AUTHOR : ISIITECH
VERSION : 0.1
// ISIITECH - Timer
// 19.01.2010 version 1.0
BEGIN

REGION Network 1 (STL): T
         A     #Input;
         JCN   ST1;
         L     #Time1;
         L     #Preset1;
         <D;
         JCN   ST2;
         A     #Pulse;
         JCN   ST2;
         L     #Time1;
         L     #Tbase;
         +D;
         T     #Time1;
         JU    ST2;
   ST1:  NOP   0;
   ST2:  NOP   0;



         A(;
         A     #RTZ;
         A     #Input_RTZ;
         );
         O(;
         AN    #Input;
         AN    #RTZ;
         );
         JCN   ST3;
         L     0;
         T     #Time1;
   ST3:  NOP   0;
END_REGION

REGION Network 2 (STL): T
         A     #Input;
         JCN   ST21;
         L     #Time2;
         L     #Preset2;
         <D;
         JCN   ST22;
         A     "point1secPls";
         JCN   ST22;
         L     #Time2;
         L     DINT#100;
         +D;
         T     #Time2;
         JU    ST22;
   ST21: NOP   0;
   ST22: NOP   0;



         A(;
         A     #RTZ;
         A     #Input_RTZ;
         );
         O(;
         AN    #Input;
         AN    #RTZ;
         );
         JCN   ST23;
         L     0;
         T     #Time2;
   ST23: NOP   0;
END_REGION
END_FUNCTION

FUNCTION "INST_CONTROL_HEATER" : Void   // FC413, LAD
TITLE = Heater controllers
{ S7_Optimized_Access := 'FALSE' }
AUTHOR : KG
VERSION : 0.1
BEGIN

REGION Network 1 (STL): Init variables
   // Dewar, Electrical Heater
         L     500.0;
         T     #Unused_TT;
         R     #ExtCmd;
END_REGION

REGION Network 2 (STL): EH90 - VB channel 1
   // Dewar, Electrical Heater
         L     2;
         T     "#DATA_HEATERS".EH90.P_TS_Ton;
         T     "#DATA_HEATERS".EH90.P_Pilot_Ton;
         L     5;
         T     "#DATA_HEATERS".EH90.P_TS_Toff;

         SET;
         A     "IOC2PLC".TT900_VALID;
         A     "EPICS_COMM_OK";
         =     #TS;
         L     "IOC2PLC".TT900;
         T     #TA;

         A(;
         L     #TA;
         L     400.0;
         >D;
         );
         JCN   _01;
         L     73.0;
         T     #TA;
   _01:  CALL  "#FC_CONTROL_HEATER"
         ( TtA      := #TA,
           TtB      := #Unused_TT,
           TtC      := #Unused_TT,
           TtD      := #Unused_TT,
           TtE      := #Unused_TT,
           TtF      := #Unused_TT,
           Nb_Tt    := 1,
           TS       := #TS,
           ExtCmd   := #ExtCmd,
           cmdEpics := "Epics_to_PLC".EH90,
           EH       := "voie 1 chaufferette BV",
           sEpics   := "PLC_to_Epics".EH90,
           Object   := "#DATA_HEATERS".EH90
         );
END_REGION

REGION Network 3 (STL): EH93-96 - VB channel 2
   // Dewar, Electrical Heater
         L     2;
         T     "#DATA_HEATERS"."EH93-96".P_TS_Ton;
         T     "#DATA_HEATERS"."EH93-96".P_Pilot_Ton;
         L     5;
         T     "#DATA_HEATERS"."EH93-96".P_TS_Toff;

         SET;
         A     "IOC2PLC".TT930_VALID;
         A     "IOC2PLC".TT940_VALID;
         A     "IOC2PLC".TT950_VALID;
         A     "IOC2PLC".TT960_VALID;
         A     "EPICS_COMM_OK";
         =     #TS;

         L     "IOC2PLC".TT930;
         T     #TA;
         A(;
         L     #TA;
         L     400.0;
         >D;
         );
         JCN   _02;
         L     73.0;
         T     #TA;
   _02:  L     "IOC2PLC".TT940;
         T     #TB;
         A(;
         L     #TB;
         L     400.0;
         >D;
         );
         JCN   _03;
         L     73.0;
         T     #TB;
   _03:  L     "IOC2PLC".TT950;
         T     #TC;
         A(;
         L     #TC;
         L     400.0;
         >D;
         );
         JCN   _04;
         L     73.0;
         T     #TC;
   _04:  L     "IOC2PLC".TT960;
         T     #TD;
         A(;
         L     #TD;
         L     400.0;
         >D;
         );
         JCN   _05;
         L     73.0;
         T     #TD;
   _05:  CALL  "#FC_CONTROL_HEATER"
         ( TtA      := #TA,
           TtB      := #TB,
           TtC      := #TC,
           TtD      := #TD,
           TtE      := #Unused_TT,
           TtF      := #Unused_TT,
           Nb_Tt    := 4,
           TS       := #TS,
           ExtCmd   := #ExtCmd,
           cmdEpics := "Epics_to_PLC"."EH93-96",
           EH       := "voie 2 chaufferette BV",
           sEpics   := "PLC_to_Epics"."EH93-96",
           Object   := "#DATA_HEATERS"."EH93-96"
         );
END_REGION

REGION Network 4 (STL): EH63_64_70 - VB channel 3
   // Dewar, Electrical Heater
         L     2;
         T     "#DATA_HEATERS"."EH63-70".P_TS_Ton;


         T     "#DATA_HEATERS"."EH63-70".P_Pilot_Ton;
         L     5;
         T     "#DATA_HEATERS"."EH63-70".P_TS_Toff;

         SET;
         A     "IOC2PLC".TT630_VALID;
         A     "IOC2PLC".TT640_VALID;
         A     "IOC2PLC".TT700_VALID;
         A     "EPICS_COMM_OK";
         =     #TS;

         CALL  "#FC_CONTROL_HEATER"
         ( TtA      := "IOC2PLC".TT630,
           TtB      := "IOC2PLC".TT640,
           TtC      := "IOC2PLC".TT700,
           TtD      := #Unused_TT,
           TtE      := #Unused_TT,
           TtF      := #Unused_TT,
           Nb_Tt    := 3,
           TS       := #TS,
           ExtCmd   := #ExtCmd,
           cmdEpics := "Epics_to_PLC"."EH63-70",
           EH       := "voie 3 chaufferette BV",
           sEpics   := "PLC_to_Epics"."EH63-70",
           Object   := "#DATA_HEATERS"."EH63-70"
         );
END_REGION

REGION Network 5 (STL): EH61-62 - VB channel 4
   // Dewar, Electrical Heater
         L     2;
         T     "#DATA_HEATERS"."EH61-62".P_TS_Ton;


         T     "#DATA_HEATERS"."EH61-62".P_Pilot_Ton;
         L     5;
         T     "#DATA_HEATERS"."EH61-62".P_TS_Toff;

         SET;
         A     "IOC2PLC".TT610_VALID;
         A     "IOC2PLC".TT620_VALID;
         A     "EPICS_COMM_OK";
         =     #TS;

         CALL  "#FC_CONTROL_HEATER"
         ( TtA      := "IOC2PLC".TT610,
           TtB      := "IOC2PLC".TT620,
           TtC      := #Unused_TT,
           TtD      := #Unused_TT,
           TtE      := #Unused_TT,
           TtF      := #Unused_TT,
           Nb_Tt    := 2,
           TS       := #TS,
           ExtCmd   := #ExtCmd,
           cmdEpics := "Epics_to_PLC"."EH61-62",
           EH       := "voie 4 chaufferette BV",
           sEpics   := "PLC_to_Epics"."EH61-62",
           Object   := "#DATA_HEATERS"."EH61-62"
         );
END_REGION

REGION Network 6 (STL): EH60_67-69 - VB channel 5
   // Dewar, Electrical Heater
         L     2;
         T     "#DATA_HEATERS"."EH60_67-69".P_TS_Ton;


         T     "#DATA_HEATERS"."EH60_67-69".P_Pilot_Ton;
         L     5;
         T     "#DATA_HEATERS"."EH60_67-69".P_TS_Toff;

         SET;
         A     "IOC2PLC".TT600_VALID;
         A     "IOC2PLC".TT670_VALID;
         A     "IOC2PLC".TT680_VALID;
         A     "IOC2PLC".TT690_VALID;
         A     "EPICS_COMM_OK";
         =     #TS;

         CALL  "#FC_CONTROL_HEATER"
         ( TtA      := "IOC2PLC".TT600,
           TtB      := "IOC2PLC".TT670,
           TtC      := "IOC2PLC".TT680,
           TtD      := "IOC2PLC".TT690,
           TtE      := #Unused_TT,
           TtF      := #Unused_TT,
           Nb_Tt    := 4,
           TS       := #TS,
           ExtCmd   := #ExtCmd,
           cmdEpics := "Epics_to_PLC"."EH60_67-69",
           EH       := "voie 5 chaufferette BV",
           sEpics   := "PLC_to_Epics"."EH60_67-69",
           Object   := "#DATA_HEATERS"."EH60_67-69"
         );
END_REGION

REGION Network 7 (STL): EH97-98 - VB channel 6
   // Dewar, Electrical Heater
         L     2;
         T     "#DATA_HEATERS"."EH97-98".P_TS_Ton;
         T     "#DATA_HEATERS"."EH97-98".P_Pilot_Ton;
         L     5;
         T     "#DATA_HEATERS"."EH97-98".P_TS_Toff;

         SET;
         A     "IOC2PLC".TT970_VALID;
         A     "IOC2PLC".TT980_VALID;
         A     "EPICS_COMM_OK";
         =     #TS;

         L     "IOC2PLC".TT970;
         T     #TA;
         A(;
         L     #TA;
         L     400.0;
         >D;
         );
         JCN   _61;
         L     73.0;
         T     #TA;
   _61:  L     "IOC2PLC".TT980;
         T     #TB;
         A(;
         L     #TB;
         L     400.0;
         >D;
         );
         JCN   _62;
         L     73.0;
         T     #TB;

   _62:  CALL  "#FC_CONTROL_HEATER"
         ( TtA      := #TA,
           TtB      := #TB,
           TtC      := #Unused_TT,
           TtD      := #Unused_TT,
           TtE      := #Unused_TT,
           TtF      := #Unused_TT,
           Nb_Tt    := 2,
           TS       := #TS,
           ExtCmd   := #ExtCmd,
           cmdEpics := "Epics_to_PLC"."EH97-98",
           EH       := "voie 6 chaufferette BV",
           sEpics   := "PLC_to_Epics"."EH97-98",
           Object   := "#DATA_HEATERS"."EH97-98"
         );
END_REGION

REGION Network 8 (STL): EH903 - CM channel 2
   // Dewar, Electrical Heater
         L     2;
         T     "#DATA_HEATERS".EH903.P_TS_Ton;
         T     "#DATA_HEATERS".EH903.P_Pilot_Ton;
         L     5;
         T     "#DATA_HEATERS".EH903.P_TS_Toff;

         SET;
         A     "IOC2PLC".TT903_VALID;
         A     "EPICS_COMM_OK";
         =     #TS;

         L     "IOC2PLC".TT903;
         T     #TA;
         A(;
         L     #TA;
         L     400.0;
         >D;
         );
         JCN   _121;
         L     73.0;
         T     #TA;
   _121: CALL  "#FC_CONTROL_HEATER"
         ( TtA      := #TA,
           TtB      := #Unused_TT,
           TtC      := #Unused_TT,
           TtD      := #Unused_TT,
           TtE      := #Unused_TT,
           TtF      := #Unused_TT,
           Nb_Tt    := 1,
           TS       := #TS,
           ExtCmd   := #ExtCmd,
           cmdEpics := "Epics_to_PLC".EH903,
           EH       := "voie 2 chaufferette CM",
           sEpics   := "PLC_to_Epics".EH903,
           Object   := "#DATA_HEATERS".EH903
         );
END_REGION

REGION Network 9 (STL): EH920 - CM channel 3
   // Dewar, Electrical Heater
         L     2;
         T     "#DATA_HEATERS".EH920.P_TS_Ton;
         T     "#DATA_HEATERS".EH920.P_Pilot_Ton;
         L     5;
         T     "#DATA_HEATERS".EH920.P_TS_Toff;

         SET;
         A     "IOC2PLC".TT920_CM_VALID;
         A     "EPICS_COMM_OK";
         =     #TS;

         L     "IOC2PLC".TT920_CM;
         T     #TA;
         A(;
         L     #TA;
         L     400.0;
         >D;
         );
         JCN   _131;
         L     73.0;
         T     #TA;
   _131: CALL  "#FC_CONTROL_HEATER"
         ( TtA      := #TA,
           TtB      := #Unused_TT,
           TtC      := #Unused_TT,
           TtD      := #Unused_TT,
           TtE      := #Unused_TT,
           TtF      := #Unused_TT,
           Nb_Tt    := 1,
           TS       := #TS,
           ExtCmd   := #ExtCmd,
           cmdEpics := "Epics_to_PLC".EH920,
           EH       := "voie 3 chaufferette CM",
           sEpics   := "PLC_to_Epics".EH920,
           Object   := "#DATA_HEATERS".EH920
         );
END_REGION

REGION Network 10 (STL): EH918 - CM channel 9
   // Dewar, Electrical Heater
         L     2;
         T     "#DATA_HEATERS".EH918.P_TS_Ton;
         T     "#DATA_HEATERS".EH918.P_Pilot_Ton;
         L     5;
         T     "#DATA_HEATERS".EH918.P_TS_Toff;

         SET;
         A     "IOC2PLC".TT918_VALID;
         A     "EPICS_COMM_OK";
         =     #TS;

         L     "IOC2PLC".TT918;
         T     #TA;
         A(;
         L     #TA;
         L     400.0;
         >D;
         );
         JCN   _191;
         L     73.0;
         T     #TA;
   _191: CALL  "#FC_CONTROL_HEATER"
         ( TtA      := #TA,
           TtB      := #Unused_TT,
           TtC      := #Unused_TT,
           TtD      := #Unused_TT,
           TtE      := #Unused_TT,
           TtF      := #Unused_TT,
           Nb_Tt    := 1,
           TS       := #TS,
           ExtCmd   := #ExtCmd,
           cmdEpics := "Epics_to_PLC".EH918,
           EH       := "voie 9 chaufferette CM",
           sEpics   := "PLC_to_Epics".EH918,
           Object   := "#DATA_HEATERS".EH918
         );
END_REGION

REGION Network 11 (STL): EH904 - CM channel 11
   // Dewar, Electrical Heater
         L     2;
         T     "#DATA_HEATERS".EH904.P_TS_Ton;
         T     "#DATA_HEATERS".EH904.P_Pilot_Ton;
         L     5;
         T     "#DATA_HEATERS".EH904.P_TS_Toff;

         SET;
         A     "IOC2PLC".TT904_VALID;
         A     "EPICS_COMM_OK";
         =     #TS;

         L     "IOC2PLC".TT904;
         T     #TA;
         A(;
         L     #TA;
         L     400.0;
         >D;
         );
         JCN   _1111;
         L     73.0;
         T     #TA;
   _1111:CALL  "#FC_CONTROL_HEATER"
         ( TtA      := #TA,
           TtB      := #Unused_TT,
           TtC      := #Unused_TT,
           TtD      := #Unused_TT,
           TtE      := #Unused_TT,
           TtF      := #Unused_TT,
           Nb_Tt    := 1,
           TS       := #TS,
           ExtCmd   := #ExtCmd,
           cmdEpics := "Epics_to_PLC".EH904,
           EH       := "voie 11 chaufferette CM",
           sEpics   := "PLC_to_Epics".EH904,
           Object   := "#DATA_HEATERS".EH904
         );
END_REGION

REGION Network 12 (STL): EH13 - Coupler 1 flange
   // Dewar, Electrical Heater
         L     2;
         T     "#DATA_HEATERS".EH13.P_TS_Ton;
         T     "#DATA_HEATERS".EH13.P_Pilot_Ton;
         L     5;
         T     "#DATA_HEATERS".EH13.P_TS_Toff;

         L     "PLC_to_Epics".TT103.Visu;
         L     0;
         ==I;
         =     #Enable;
         CALL  "#FC_CONTROL_HEATER"
         ( TtA      := "PLC_to_Epics".TT103.Level,
           TtB      := #Unused_TT,
           TtC      := #Unused_TT,
           TtD      := #Unused_TT,
           TtE      := #Unused_TT,
           TtF      := #Unused_TT,
           Nb_Tt    := 1,
           TS       := #Enable,
           ExtCmd   := #ExtCmd,
           cmdEpics := "Epics_to_PLC".EH13,
           EH       := "EH13 Cpl1",
           sEpics   := "PLC_to_Epics".EH13,
           Object   := "#DATA_HEATERS".EH13
         );
END_REGION

REGION Network 13 (STL): EH43 - Coupler 2 flange
   // Dewar, Electrical Heater
         L     2;
         T     "#DATA_HEATERS".EH43.P_TS_Ton;
         T     "#DATA_HEATERS".EH43.P_Pilot_Ton;
         L     5;
         T     "#DATA_HEATERS".EH43.P_TS_Toff;

         L     "PLC_to_Epics".TT203.Visu;
         L     0;
         ==I;
         =     #Enable;
         CALL  "#FC_CONTROL_HEATER"
         ( TtA      := "PLC_to_Epics".TT203.Level,
           TtB      := #Unused_TT,
           TtC      := #Unused_TT,
           TtD      := #Unused_TT,
           TtE      := #Unused_TT,
           TtF      := #Unused_TT,
           Nb_Tt    := 1,
           TS       := #Enable,
           ExtCmd   := #ExtCmd,
           cmdEpics := "Epics_to_PLC".EH43,
           EH       := "EH43 Cpl2",
           sEpics   := "PLC_to_Epics".EH43,
           Object   := "#DATA_HEATERS".EH43
         );
END_REGION
END_FUNCTION

FUNCTION "Manage_HEATERS" : Void   // FC513, LAD
TITLE = Manage the heaters
{ S7_Optimized_Access := 'FALSE' }
AUTHOR : KG
VERSION : 0.1
BEGIN

REGION Network 1: EH13 & EH43 - Coupler flange cavity 1 and 2
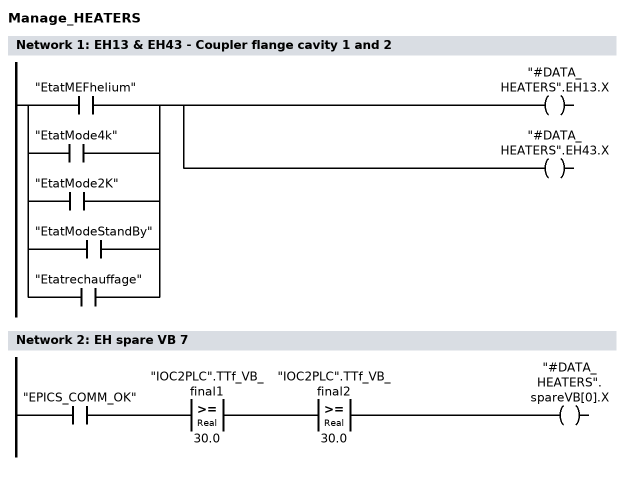
   RUNG wire#powerrail
      Contact( "EtatMEFhelium" )
      wire#w1
      Coil( "#DATA_HEATERS".EH13.X )
   END_RUNG
   RUNG wire#powerrail
      Contact( "EtatMode4k" )
   END_RUNG wire#w1
   RUNG wire#powerrail
      Contact( "EtatMode2K" )
   END_RUNG wire#w1
   RUNG wire#powerrail
      Contact( "EtatModeStandBy" )
   END_RUNG wire#w1
   RUNG wire#powerrail
      Contact( "Etatrechauffage" )
   END_RUNG wire#w1
   RUNG wire#w1
      Coil( "#DATA_HEATERS".EH43.X )
   END_RUNG
   // the same network as SCL:
   "#DATA_HEATERS".EH13.X := "EtatMEFhelium" OR "EtatMode4k" OR "EtatMode2K" OR "EtatModeStandBy" OR "Etatrechauffage";
   "#DATA_HEATERS".EH43.X := "#DATA_HEATERS".EH13.X;
END_REGION

REGION Network 2: EH spare VB 7
   RUNG wire#powerrail
      Contact( "EPICS_COMM_OK" )
      { S7_Templates := "SrcType := Real" } GE_Contact(in1 := "IOC2PLC".TTf_VB_final1, in2 := 30.0)
      { S7_Templates := "SrcType := Real" } GE_Contact(in1 := "IOC2PLC".TTf_VB_final2, in2 := 30.0)
      Coil( "#DATA_HEATERS".spareVB[0].X )
   END_RUNG
   // the same network as SCL:
   "#DATA_HEATERS".spareVB[0].X := "EPICS_COMM_OK" AND ("IOC2PLC".TTf_VB_final1 >= 30.0) AND ("IOC2PLC".TTf_VB_final2 >= 30.0);
END_REGION
END_FUNCTION

ORGANIZATION_BLOCK "Main"   // OB1, STL
TITLE = "Main Program Sweep (Cycle)"
{ S7_Optimized_Access := 'FALSE' }
VERSION : 0.1
BEGIN

REGION Network 1: Set-up the timing pulse for FC_TIMER
         A     "point1sec";
         AN    "point1secMem";
         =     "point1secPls";
         A     "point1sec";
         =     "point1secMem";

         SET;
         A     "oneSec";
         AN    "oneSecMem";
         =     "oneSecPls";
         A     "oneSec";
         =     "oneSecMem";
END_REGION

REGION Network 2: Get data and commands from Epics IOC
         CALL  "Recv_from_Epics";
         NOP   0;
END_REGION

REGION Network 3
         A     "Graph/manuelle";
         JNB   Label_0;
         CALL  "commande vanne";
   Label_0:NOP   0;
END_REGION

REGION Network 4
         CALL  "NIveau Helium&Pression&vide";
         NOP   0;
END_REGION

REGION Network 5
         CALL  "ACQ_CABTF";
         NOP   0;
END_REGION

REGION Network 6
         AN    "Graph/manuelle";
         JNB   Label_1;
         CALL  "grafcet";
   Label_1:NOP   0;
END_REGION

REGION Network 7
         CALL  "Send_to_Epics";
         NOP   0;
END_REGION

REGION Network 8: Instantiate the heaters control
         CALL  "INST_CONTROL_HEATER";
END_REGION

REGION Network 9: Manage the heaters
         CALL  "Manage_HEATERS";
END_REGION

REGION Network 10: Clear INIT flag after the first cycle
         SET;
         R     "INIT";
END_REGION

REGION Network 11
         CALL  "UpdateData2HNOSS";
END_REGION

REGION Network 12: Appeler le bloc de diagnostic système / Call system diagnostics block
         CALL  "RSE_FB", "RSE_DB";
END_REGION
END_ORGANIZATION_BLOCK

ORGANIZATION_BLOCK "CYC_INT2"   // OB32, LAD
TITLE = Cyclic_1s / "Cyclic Interrupt"
{ S7_Optimized_Access := 'FALSE' }
AUTHOR : KG
VERSION : 0.1
// Call the PID functionswith 1s interval
   VAR_TEMP   // added for the SCL form of the ladder/FBD networks
      _w1 : Bool;
   END_VAR
BEGIN

REGION Network 1: PID regulator for the LN2 screen cooling (CV60)
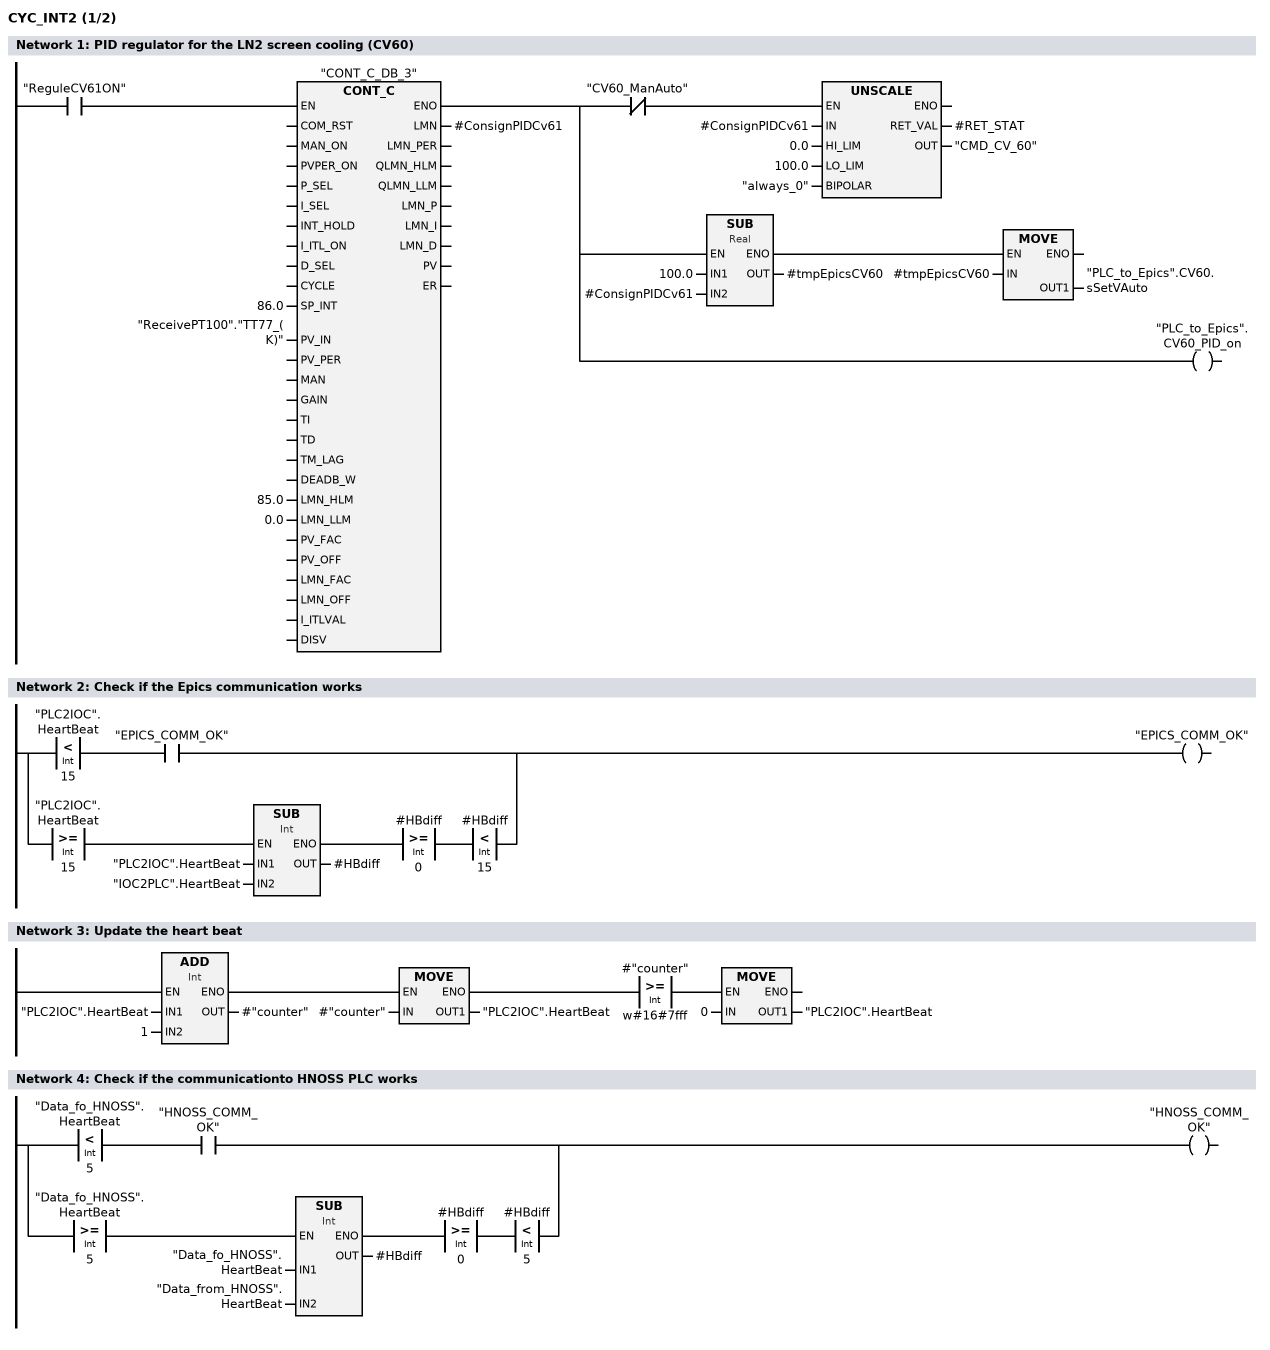
   // ENO of a box is taken as its EN; it also drops when the box reports an error
   #_w1 := "ReguleCV61ON";
   IF #_w1 THEN
       "CONT_C_DB_3"(SP_INT := 86.0,   // CONT_C
                     PV_IN := "ReceivePT100"."TT77_(K)",
                     LMN_HLM := 85.0,
                     LMN_LLM := 0.0,
                     LMN => #ConsignPIDCv61);
   END_IF;
   IF #_w1 AND NOT "CV60_ManAuto" THEN
       #RET_STAT := UNSCALE(IN := #ConsignPIDCv61,
                            HI_LIM := 0.0,
                            LO_LIM := 100.0,
                            BIPOLAR := "always_0",
                            OUT => "CMD_CV_60");
   END_IF;
   IF #_w1 THEN
       #tmpEpicsCV60 := 100.0 - #ConsignPIDCv61;
       "PLC_to_Epics".CV60.sSetVAuto := #tmpEpicsCV60;
   END_IF;
   "PLC_to_Epics".CV60_PID_on := #_w1;
END_REGION

REGION Network 2: Check if the Epics communication works
   RUNG wire#powerrail
      { S7_Templates := "SrcType := Int" } LT_Contact(in1 := "PLC2IOC".HeartBeat, in2 := 15)
      Contact( "EPICS_COMM_OK" )
      wire#w1
      Coil( "EPICS_COMM_OK" )
   END_RUNG
   RUNG wire#powerrail
      { S7_Templates := "SrcType := Int" } GE_Contact(in1 := "PLC2IOC".HeartBeat, in2 := 15)
      { S7_Templates := "SrcType := Int"; S7_GenerateENO := "TRUE" } Sub(in1 := "PLC2IOC".HeartBeat, in2 := "IOC2PLC".HeartBeat, out => #HBdiff)
      { S7_Templates := "SrcType := Int" } GE_Contact(in1 := #HBdiff, in2 := 0)
      { S7_Templates := "SrcType := Int" } LT_Contact(in1 := #HBdiff, in2 := 15)
   END_RUNG wire#w1
   // the same network as SCL:
   // ENO of a box is taken as its EN; it also drops when the box reports an error
   #_w1 := "PLC2IOC".HeartBeat >= 15;
   IF #_w1 THEN #HBdiff := "PLC2IOC".HeartBeat - "IOC2PLC".HeartBeat; END_IF;
   "EPICS_COMM_OK" := (("PLC2IOC".HeartBeat < 15) AND "EPICS_COMM_OK") OR (#_w1 AND (#HBdiff >= 0) AND (#HBdiff < 15));
END_REGION

REGION Network 3: Update the heart beat
   RUNG wire#powerrail
      { S7_Templates := "SrcType := Int"; S7_GenerateENO := "TRUE" } Add(in1 := "PLC2IOC".HeartBeat, in2 := 1, out => #"counter")
      { S7_GenerateENO := "TRUE" } Move(in := #"counter", out1 => "PLC2IOC".HeartBeat)
      { S7_Templates := "SrcType := Int" } GE_Contact(in1 := #"counter", in2 := w#16#7fff)
      { S7_GenerateENO := "TRUE" } Move(in := 0, out1 => "PLC2IOC".HeartBeat)
   END_RUNG
   // the same network as SCL:
   // ENO of a box is taken as its EN; it also drops when the box reports an error
   #"counter" := "PLC2IOC".HeartBeat + 1;
   "PLC2IOC".HeartBeat := #"counter";
   IF #"counter" >= w#16#7fff THEN "PLC2IOC".HeartBeat := 0; END_IF;
END_REGION

REGION Network 4: Check if the communicationto HNOSS PLC works
   RUNG wire#powerrail
      { S7_Templates := "SrcType := Int" } LT_Contact(in1 := "Data_fo_HNOSS".HeartBeat, in2 := 5)
      Contact( "HNOSS_COMM_OK" )
      wire#w1
      Coil( "HNOSS_COMM_OK" )
   END_RUNG
   RUNG wire#powerrail
      { S7_Templates := "SrcType := Int" } GE_Contact(in1 := "Data_fo_HNOSS".HeartBeat, in2 := 5)
      { S7_Templates := "SrcType := Int"; S7_GenerateENO := "TRUE" } Sub(in1 := "Data_fo_HNOSS".HeartBeat, in2 := "Data_from_HNOSS".HeartBeat, out => #HBdiff)
      { S7_Templates := "SrcType := Int" } GE_Contact(in1 := #HBdiff, in2 := 0)
      { S7_Templates := "SrcType := Int" } LT_Contact(in1 := #HBdiff, in2 := 5)
   END_RUNG wire#w1
   // the same network as SCL:
   // ENO of a box is taken as its EN; it also drops when the box reports an error
   #_w1 := "Data_fo_HNOSS".HeartBeat >= 5;
   IF #_w1 THEN #HBdiff := "Data_fo_HNOSS".HeartBeat - "Data_from_HNOSS".HeartBeat; END_IF;
   "HNOSS_COMM_OK" := (("Data_fo_HNOSS".HeartBeat < 5) AND "HNOSS_COMM_OK") OR (#_w1 AND (#HBdiff >= 0) AND (#HBdiff < 5));
END_REGION

REGION Network 5: Update the heart beat
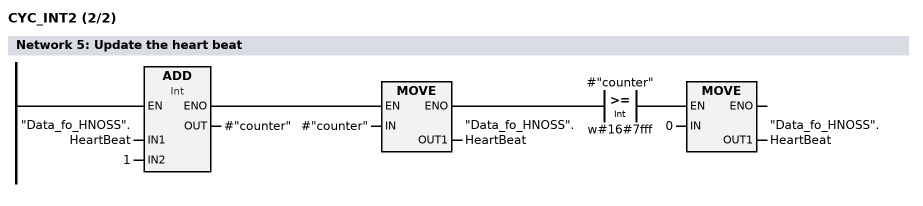
   RUNG wire#powerrail
      { S7_Templates := "SrcType := Int"; S7_GenerateENO := "TRUE" } Add(in1 := "Data_fo_HNOSS".HeartBeat, in2 := 1, out => #"counter")
      { S7_GenerateENO := "TRUE" } Move(in := #"counter", out1 => "Data_fo_HNOSS".HeartBeat)
      { S7_Templates := "SrcType := Int" } GE_Contact(in1 := #"counter", in2 := w#16#7fff)
      { S7_GenerateENO := "TRUE" } Move(in := 0, out1 => "Data_fo_HNOSS".HeartBeat)
   END_RUNG
   // the same network as SCL:
   // ENO of a box is taken as its EN; it also drops when the box reports an error
   #"counter" := "Data_fo_HNOSS".HeartBeat + 1;
   "Data_fo_HNOSS".HeartBeat := #"counter";
   IF #"counter" >= w#16#7fff THEN "Data_fo_HNOSS".HeartBeat := 0; END_IF;
END_REGION
END_ORGANIZATION_BLOCK

ORGANIZATION_BLOCK "CYC_INT5"   // OB35, LAD
TITLE = "Cyclic Interrupt"
{ S7_Optimized_Access := 'FALSE' }
VERSION : 0.1
   VAR_TEMP   // added for the SCL form of the ladder/FBD networks
      _w1 : Bool;
      _w2 : Bool;
   END_VAR
BEGIN

REGION Network 1
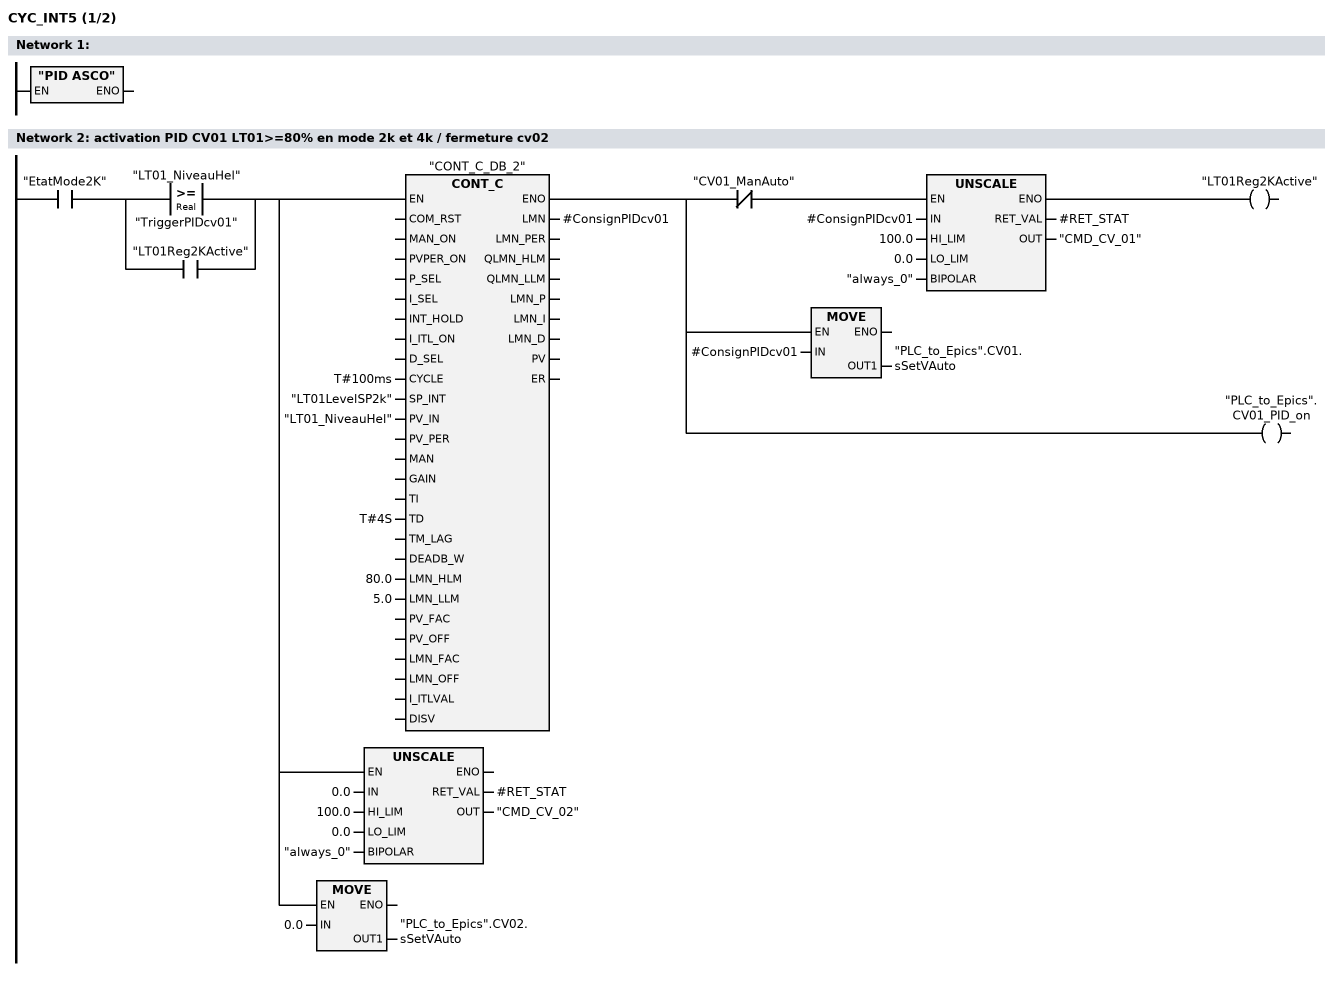
   RUNG wire#powerrail
      "PID ASCO"()
   END_RUNG
   // the same network as SCL:
   "PID ASCO"();
END_REGION

REGION Network 2: activation PID CV01 LT01>=80% en mode 2k et 4k / fermeture cv02
   // ENO of a box is taken as its EN; it also drops when the box reports an error
   #_w1 := "EtatMode2K" AND (("LT01_NiveauHel" >= "TriggerPIDcv01") OR "LT01Reg2KActive");
   IF #_w1 THEN
       "CONT_C_DB_2"(CYCLE := T#100ms,   // CONT_C
                     SP_INT := "LT01LevelSP2k",
                     PV_IN := "LT01_NiveauHel",
                     TD := T#4S,
                     LMN_HLM := 80.0,
                     LMN_LLM := 5.0,
                     LMN => #ConsignPIDcv01);
   END_IF;
   #_w2 := #_w1 AND NOT "CV01_ManAuto";
   IF #_w2 THEN
       #RET_STAT := UNSCALE(IN := #ConsignPIDcv01,
                            HI_LIM := 100.0,
                            LO_LIM := 0.0,
                            BIPOLAR := "always_0",
                            OUT => "CMD_CV_01");
   END_IF;
   "LT01Reg2KActive" := #_w2;
   IF #_w1 THEN "PLC_to_Epics".CV01.sSetVAuto := #ConsignPIDcv01; END_IF;
   "PLC_to_Epics".CV01_PID_on := #_w1;
   IF #_w1 THEN
       #RET_STAT := UNSCALE(IN := 0.0, HI_LIM := 100.0, LO_LIM := 0.0, BIPOLAR := "always_0", OUT => "CMD_CV_02");
       "PLC_to_Epics".CV02.sSetVAuto := 0.0;
   END_IF;
END_REGION

REGION Network 3: activation PID CV03 LT03>=80%
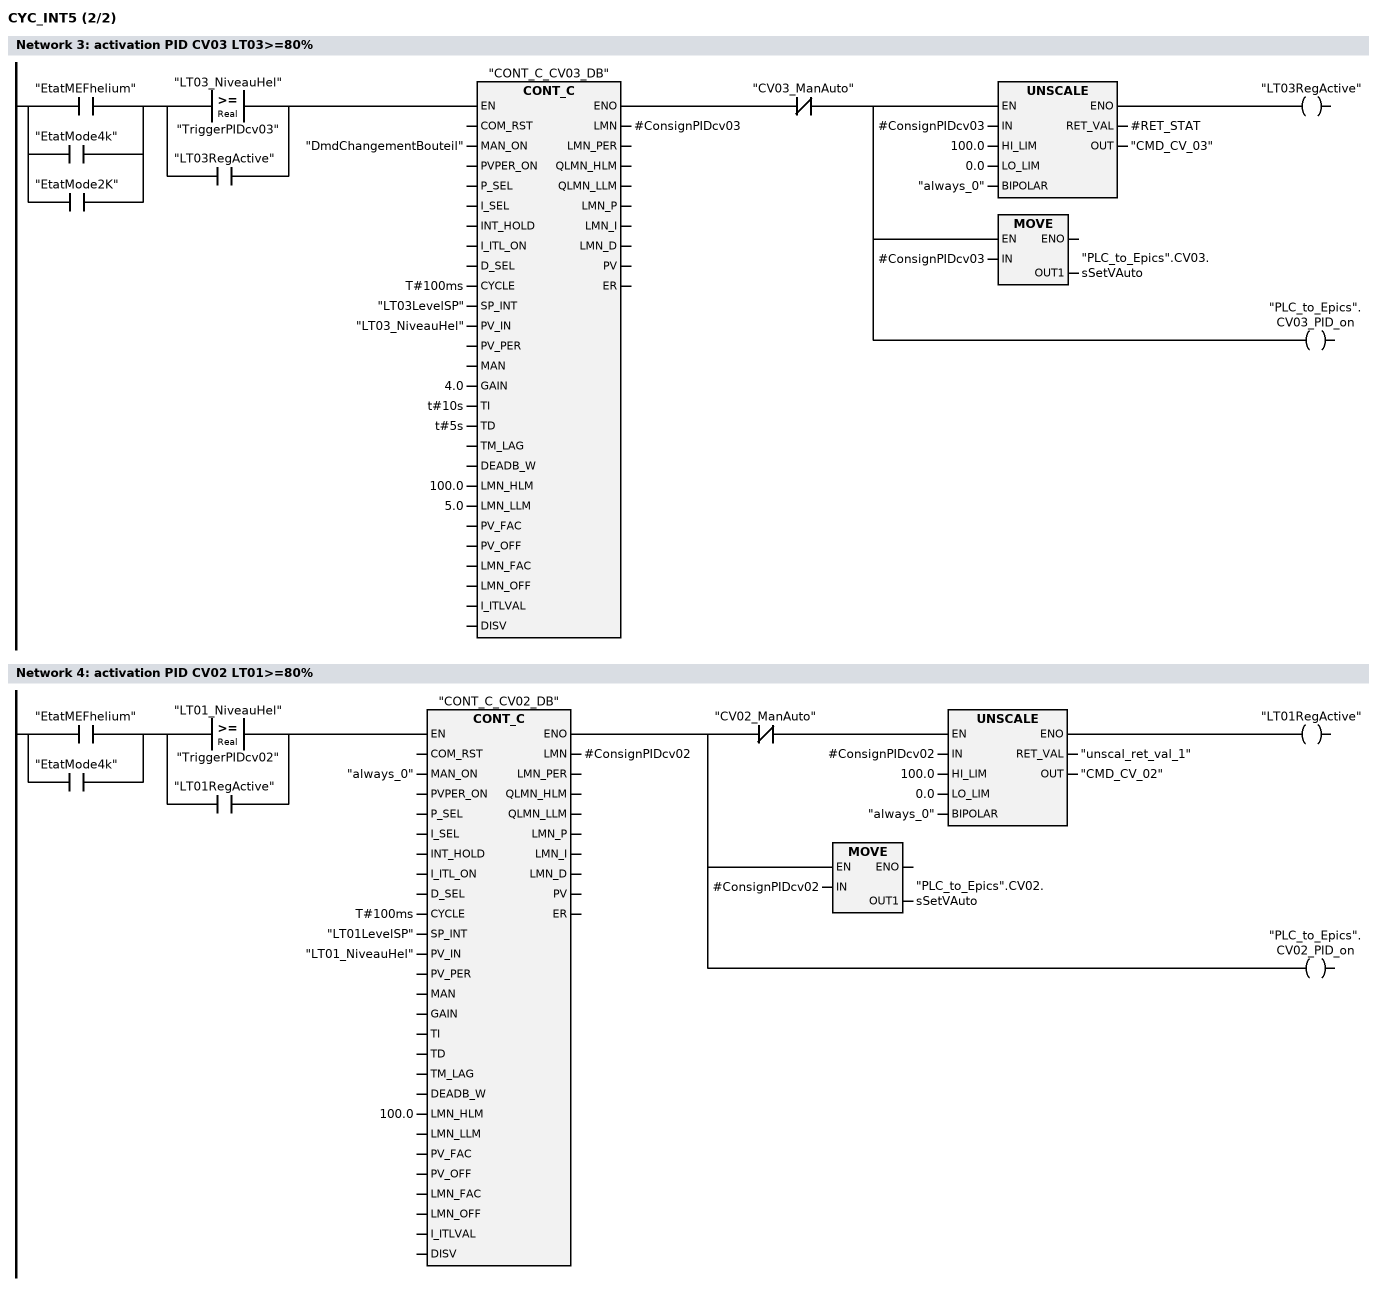
   // ENO of a box is taken as its EN; it also drops when the box reports an error
   #_w1 := ("EtatMEFhelium" OR "EtatMode4k" OR "EtatMode2K") AND (("LT03_NiveauHel" >= "TriggerPIDcv03") OR "LT03RegActive");
   IF #_w1 THEN
       "CONT_C_CV03_DB"(MAN_ON := "DmdChangementBouteil",   // CONT_C
                        CYCLE := T#100ms,
                        SP_INT := "LT03LevelSP",
                        PV_IN := "LT03_NiveauHel",
                        GAIN := 4.0,
                        TI := t#10s,
                        TD := t#5s,
                        LMN_HLM := 100.0,
                        LMN_LLM := 5.0,
                        LMN => #ConsignPIDcv03);
   END_IF;
   #_w2 := #_w1 AND NOT "CV03_ManAuto";
   IF #_w2 THEN
       #RET_STAT := UNSCALE(IN := #ConsignPIDcv03,
                            HI_LIM := 100.0,
                            LO_LIM := 0.0,
                            BIPOLAR := "always_0",
                            OUT => "CMD_CV_03");
   END_IF;
   "LT03RegActive" := #_w2;
   IF #_w2 THEN "PLC_to_Epics".CV03.sSetVAuto := #ConsignPIDcv03; END_IF;
   "PLC_to_Epics".CV03_PID_on := #_w2;
END_REGION

REGION Network 4: activation PID CV02 LT01>=80%
   // ENO of a box is taken as its EN; it also drops when the box reports an error
   #_w1 := ("EtatMEFhelium" OR "EtatMode4k") AND (("LT01_NiveauHel" >= "TriggerPIDcv02") OR "LT01RegActive");
   IF #_w1 THEN
       "CONT_C_CV02_DB"(MAN_ON := "always_0",   // CONT_C
                        CYCLE := T#100ms,
                        SP_INT := "LT01LevelSP",
                        PV_IN := "LT01_NiveauHel",
                        LMN_HLM := 100.0,
                        LMN => #ConsignPIDcv02);
   END_IF;
   #_w2 := #_w1 AND NOT "CV02_ManAuto";
   IF #_w2 THEN
       "unscal_ret_val_1" := UNSCALE(IN := #ConsignPIDcv02,
                               HI_LIM := 100.0,
                               LO_LIM := 0.0,
                               BIPOLAR := "always_0",
                               OUT => "CMD_CV_02");
   END_IF;
   "LT01RegActive" := #_w2;
   IF #_w1 THEN "PLC_to_Epics".CV02.sSetVAuto := #ConsignPIDcv02; END_IF;
   "PLC_to_Epics".CV02_PID_on := #_w1;
END_REGION
END_ORGANIZATION_BLOCK

ORGANIZATION_BLOCK "HW_INT0"   // OB40, LAD
TITLE = "Hardware Interrupt"
{ S7_Optimized_Access := 'FALSE' }
VERSION : 0.1
BEGIN
END_ORGANIZATION_BLOCK

ORGANIZATION_BLOCK "I/O_FLT1"   // OB82, LAD
TITLE = "I/O Point Fault"
{ S7_Optimized_Access := 'FALSE' }
VERSION : 0.1
BEGIN

REGION Network 1 (STL): Appeler le bloc de diagnostic système / Call system diagnostics block
         CALL  "RSE_FB", "RSE_DB";
END_REGION
END_ORGANIZATION_BLOCK

ORGANIZATION_BLOCK "OBNL_FLT"   // OB85, LAD
TITLE = "Organization Block (OB) Not Loaded Fault"
{ S7_Optimized_Access := 'FALSE' }
VERSION : 0.1
BEGIN
END_ORGANIZATION_BLOCK

ORGANIZATION_BLOCK "RACK_FLT"   // OB86, LAD
TITLE = "Loss Of Rack Fault"
{ S7_Optimized_Access := 'FALSE' }
VERSION : 0.1
BEGIN

REGION Network 1 (STL): Appeler le bloc de diagnostic système / Call system diagnostics block
         CALL  "RSE_FB", "RSE_DB";
END_REGION
END_ORGANIZATION_BLOCK

ORGANIZATION_BLOCK "COMPLETE RESTART"   // OB100, STL
TITLE = "Complete Restart"
{ S7_Optimized_Access := 'FALSE' }
VERSION : 0.1
BEGIN

REGION Network 1
         SET;
         S     "INIT";
END_REGION
END_ORGANIZATION_BLOCK

(* ===== HMI "HMI_RT_1" =====

graphic list "Vanne horizontale maxi_0": 1 'Vanne horizontale verte_2'; 0 'Vanne horizontale rouge_2'; 2 'Vanne horizontale rouge_2'; 3 'Vanne horizontale verte_2'; 4 'Vanne horizontale grise_2'; 5 'Vanne horizontale grise_2'

ScreenModuleEditorView "Bloc Vanne horizontale" 1024x768
   GraphicIOField "Modèle_Champ E/S graphique_13" at 10,10 size 50x35
*)

(* ===== HMI "HMI_RT_1" =====

graphic list "Vanne verticale maxi_0": 1 'Vanne verticale verte_1'; 2 'Vanne verticale rouge_1'; 0 'Vanne verticale rouge_1'; 3 'Vanne verticale verte_1'; 4 'Vanne verticale grise_1'; 5 'Vanne verticale grise_1'

ScreenModuleEditorView "Bloc Vanne verticale" 1024x768
   GraphicIOField "Champ E/S graphique_10" at 10,10 size 35x50
*)